HMI tags "IGG import"
   "RESET_STEP" : Bool = PLC RESET_STEP AT %M12.0, 1 s
   "Start Sequenc_DB_Post Purge Time Sec" : Int AT %DB1.DBW0
   "Tank Activated Port 10" : Int AT %DB1.DBW0
   "Tank Activated Port 2" : Int AT %DB1.DBW0
   "Tank Activated Port 3" : Int AT %DB1.DBW0
   "Tank Activated Port 4" : Int AT %DB1.DBW0
   "Tank Activated Port 5" : Int AT %DB1.DBW0
   "Tank Activated Port 6" : Int AT %DB1.DBW0
   "Tank Activated Port 7" : Int AT %DB1.DBW0
   "Tank Activated Port 8" : Int AT %DB1.DBW0
   "Tank Activated Port 9" : Int AT %DB1.DBW0
   "Tank Activated Star 10" : Int AT %DB1.DBW0
   "Tank Activated Star 2" : Int AT %DB1.DBW0
   "Tank Activated Star 3" : Int AT %DB1.DBW0
   "Tank Activated Star 4" : Int AT %DB1.DBW0
   "Tank Activated Star 5" : Int AT %DB1.DBW0
   "Tank Activated Star 6" : Int AT %DB1.DBW0
   "Tank Activated Star 7" : Int AT %DB1.DBW0
   "Tank Activated Star 8" : Int AT %DB1.DBW0
   "Tank Activated Star 9" : Int AT %DB1.DBW0
   "user_group" : Int AT %DB1.DBW0
   "2084_Setpoints_FIT417_HiHi" : Real = PLC "2084_Setpoints".FIT417_HiHi, 1 s
   "2086_Times_Tank Alarm Reset Time" : Time = PLC "2086_Times"."Tank Alarm Reset Time", 1 s
   "2084_Setpoints_FIT417_LoLo" : Real = PLC "2084_Setpoints".FIT417_LoLo, 1 s
   "2086_Times_Alarm Enable Delay" : Time = PLC "2086_Times"."Alarm Enable Delay", 1 s
   "2084_Setpoints_FIT417_Lo" : Real = PLC "2084_Setpoints".FIT417_Lo, 1 s
   "2084_Setpoints_FIT419_Lo" : Real = PLC "2084_Setpoints".FIT419_Lo, 1 s
   "2084_Setpoints_FIT417_Hi" : Real = PLC "2084_Setpoints".FIT417_Hi, 1 s
   "LT422 FPT  TANK LEVEL ALARM_LOW LEVEL VALUE (L)" : Real = PLC "LT422 FPT  TANK LEVEL ALARM"."LOW LEVEL VALUE (L)" AT %DB2226.DBD26, 1 s
   "2084_Setpoints_FIT419_LoLo" : Real = PLC "2084_Setpoints".FIT419_LoLo, 1 s
   "LT422 FPT  TANK LEVEL ALARM_ALARM L" : Bool = PLC "LT422 FPT  TANK LEVEL ALARM"."ALARM L" AT %DB2226.DBX48.2, 1 s
   "20_TANKS_IP_DATA_RIO_03_FIRST_TANK_O2_MONITOR" : Real = PLC "20_TANKS_IP_DATA".RIO_03.FIRST_TANK.O2_MONITOR, 1 s
   "20_TANKS_IP_DATA_RIO_07_FIRST_TANK_DECK_IG_PRESS" : Real = PLC "20_TANKS_IP_DATA".RIO_07.FIRST_TANK.DECK_IG_PRESS, 1 s
   "2062_Warning_Data_Alarm Tank FPT" : Bool = PLC "2062_Warning_Data"."Alarm Tank FPT" AT %DB2062.DBX22.1, 1 s
   "2084_Setpoints_LT421_Hi" : Real = PLC "2084_Setpoints".LT421_Hi, 1 s
   "2084_Setpoints_TX426 Port PH Lo" : Real = PLC "2084_Setpoints"."TX426 Port PH Lo", 1 s
   "2084_Setpoints_TX426 Port PH High" : Real = PLC "2084_Setpoints"."TX426 Port PH High", 1 s
   "2084_Setpoints_TX428 Port DO Lo" : Real = PLC "2084_Setpoints"."TX428 Port DO Lo", 1 s
   "2084_Setpoints_TX428 Port DO High" : Real = PLC "2084_Setpoints"."TX428 Port DO High", 1 s
   "2084_Setpoints_LT421_Lo" : Real = PLC "2084_Setpoints".LT421_Lo, 1 s
   "2084_Setpoints_FIT419_HiHi" : Real = PLC "2084_Setpoints".FIT419_HiHi, 1 s
   "2084_Setpoints_FIT419_Hi" : Real = PLC "2084_Setpoints".FIT419_Hi, 1 s
   "2084_Setpoints_TX425 Star PH Lo" : Real = PLC "2084_Setpoints"."TX425 Star PH Lo", 1 s
   "2084_Setpoints_TX425 Star PH High" : Real = PLC "2084_Setpoints"."TX425 Star PH High", 1 s
   "2084_Setpoints_TX427 Star DO Lo" : Real = PLC "2084_Setpoints"."TX427 Star DO Lo", 1 s
   "2084_Setpoints_TX427 Star DO High" : Real = PLC "2084_Setpoints"."TX427 Star DO High", 1 s
   "2084_Setpoints_Conf O2 Level Lo" : Real = PLC "2084_Setpoints"."Conf O2 Level Lo", 1 s
   "2084_Setpoints_Conf O2 Level Lo Lo" : Real = PLC "2084_Setpoints"."Conf O2 Level Lo Lo", 1 s
   "20_TANKS_IP_DATA_RIO_03_FIRST_TANK_DECK_IG_PRESS" : Real = PLC "20_TANKS_IP_DATA".RIO_03.FIRST_TANK.DECK_IG_PRESS, 1 s
   "20_TANKS_IP_DATA_RIO_01_THIRD_TANK_O2_MONITOR" : Real = PLC "20_TANKS_IP_DATA".RIO_01.THIRD_TANK.O2_MONITOR, 1 s
   "20_TANKS_IP_DATA_RIO_01_THIRD_TANK_DECK_IG_PRESS" : Real = PLC "20_TANKS_IP_DATA".RIO_01.THIRD_TANK.DECK_IG_PRESS, 1 s
   "20_TANKS_IP_DATA_RIO_01_FIRST_TANK_DECK_IG_PRESS" : Real = PLC "20_TANKS_IP_DATA".RIO_01.FIRST_TANK.DECK_IG_PRESS, 1 s
   "20_TANKS_IP_DATA_RIO_01_FIRST_TANK_O2_MONITOR" : Real = PLC "20_TANKS_IP_DATA".RIO_01.FIRST_TANK.O2_MONITOR, 1 s
   "20_TANKS_IP_DATA_RIO_04_FIRST_TANK_DECK_IG_PRESS" : Real = PLC "20_TANKS_IP_DATA".RIO_04.FIRST_TANK.DECK_IG_PRESS, 1 s
   "20_TANKS_IP_DATA_RIO_04_FIRST_TANK_O2_MONITOR" : Real = PLC "20_TANKS_IP_DATA".RIO_04.FIRST_TANK.O2_MONITOR, 1 s
   "20_TANKS_IP_DATA_RIO_04_SECOND_TANK_O2_MONITOR" : Real = PLC "20_TANKS_IP_DATA".RIO_04.SECOND_TANK.O2_MONITOR, 1 s
   "20_TANKS_IP_DATA_RIO_05_FIRST_TANK_DECK_IG_PRESS" : Real = PLC "20_TANKS_IP_DATA".RIO_05.FIRST_TANK.DECK_IG_PRESS, 1 s
   "20_TANKS_IP_DATA_RIO_05_FIRST_TANK_O2_MONITOR" : Real = PLC "20_TANKS_IP_DATA".RIO_05.FIRST_TANK.O2_MONITOR, 1 s
   "20_TANKS_IP_DATA_RIO_05_SECOND_TANK_O2_MONITOR" : Real = PLC "20_TANKS_IP_DATA".RIO_05.SECOND_TANK.O2_MONITOR, 1 s
   "20_TANKS_IP_DATA_RIO_06_FIRST_TANK_DECK_IG_PRESS" : Real = PLC "20_TANKS_IP_DATA".RIO_06.FIRST_TANK.DECK_IG_PRESS, 1 s
   "20_TANKS_IP_DATA_RIO_06_FIRST_TANK_O2_MONITOR" : Real = PLC "20_TANKS_IP_DATA".RIO_06.FIRST_TANK.O2_MONITOR, 1 s
   "20_TANKS_IP_DATA_RIO_07_FIRST_TANK_O2_MONITOR" : Real = PLC "20_TANKS_IP_DATA".RIO_07.FIRST_TANK.O2_MONITOR, 1 s
   "20_TANKS_IP_DATA_RIO_03_SECOND_TANK_O2_MONITOR" : Real = PLC "20_TANKS_IP_DATA".RIO_03.SECOND_TANK.O2_MONITOR, 1 s
   "2062_Warning_Data_Water Level Override FPT" : Bool = PLC "2062_Warning_Data"."Water Level Override FPT" AT %DB2062.DBX360.0, 1 s
   "Tank 3P Tank Vent Valve 2 Feedback - Closed" : Bool = PLC "Tank 3P Tank Vent Valve 2 Feedback - Closed" AT %I27.5, 1 s
   "2062_Warning_Data_Alarm Tank P1" : Bool = PLC "2062_Warning_Data"."Alarm Tank P1" AT %DB2062.DBX22.2, 1 s
   "Tank 2S Tank Vent Valve 2 Feedback - Opened" : Bool = PLC "Tank 2S Tank Vent Valve 2 Feedback - Opened" AT %I18.4, 1 s
   "Tank 2S Tank Vent Valve 1 Feedback - Closed" : Bool = PLC "Tank 2S Tank Vent Valve 1 Feedback - Closed" AT %I18.3, 1 s
   "Tank 2S Tank Vent Valve 1 Feedback - Opened" : Bool = PLC "Tank 2S Tank Vent Valve 1 Feedback - Opened" AT %I18.2, 1 s
   "Tank 2S GTT Isolation Valve Feedback - Closed" : Bool = PLC "Tank 2S GTT Isolation Valve Feedback - Closed" AT %I18.1, 1 s
   "Tank 2S GTT Isolation Valve Feedback - Opened" : Bool = PLC "Tank 2S GTT Isolation Valve Feedback - Opened" AT %I18.0, 1 s
   "RIO2_SPR_DI_15_7" : Bool = PLC RIO2_SPR_DI_15_7 AT %I15.7, 1 s
   "RIO2_SPR_DI_15_6" : Bool = PLC RIO2_SPR_DI_15_6 AT %I15.6, 1 s
   "Tank 2P Tank Vent Valve 2 Feedback - Closed" : Bool = PLC "20_TANKS_IP_DATA".RIO_05.FIRST_TANK.BWT_DO AT %I15.5, 1 s
   "Tank 2P Tank Vent Valve 2 Feedback - Opened" : Bool = PLC "Tank 2P Tank Vent Valve 2 Feedback - Opened" AT %I15.4, 1 s
   "Tank 2P Tank Vent Valve 1 Feedback - Closed" : Bool = PLC "Tank 2P Tank Vent Valve 1 Feedback - Closed" AT %I15.3, 1 s
   "Tank 2P Tank Vent Valve 1 Feedback - Opened" : Bool = PLC "Tank 2P Tank Vent Valve 1 Feedback - Opened" AT %I15.2, 1 s
   "Tank 2S Tank Vent Valve 2 Feedback - Closed" : Bool = PLC "Tank 2S Tank Vent Valve 2 Feedback - Closed" AT %I18.5, 1 s
   "Tank 2P GTT Isolation Valve Feedback - Closed" : Bool = PLC "Tank 2P GTT Isolation Valve Feedback - Closed" AT %I15.1, 1 s
   "RIO1_SPR_DI_9_7" : Bool = PLC RIO1_SPR_DI_9_7 AT %I9.7, 1 s
   "RIO1_SPR_DI_9_6" : Bool = PLC RIO1_SPR_DI_9_6 AT %I9.6, 1 s
   "RIO1_SPR_DI_9_5" : Bool = PLC RIO1_SPR_DI_9_5 AT %I9.5, 1 s
   "RIO1_SPR_DI_9_4" : Bool = PLC RIO1_SPR_DI_9_4 AT %I9.4, 1 s
   "Tank 1S BWT Level High High Switch" : Bool = PLC "Tank 1S BWT Level High High Switch" AT %I9.3, 1 s
   "Tank 1P BWT Level High High Switch" : Bool = PLC "Tank 1P BWT Level High High Switch" AT %I9.2, 1 s
   "RIO1 Tanks Pressure Switch Hi Hi" : Bool = PLC "RIO1 Tanks Pressure Switch Hi Hi" AT %I9.1, 1 s
   "FPT BWT Level High High Switch" : Bool = PLC "FPT BWT Level High High Switch" AT %I9.0, 1 s
   "RIO1_SPR_DI_6_7" : Bool = PLC RIO1_SPR_DI_6_7 AT %I6.7, 1 s
   "RIO1_SPR_DI_6_6" : Bool = PLC RIO1_SPR_DI_6_6 AT %I6.6, 1 s
   "Tank 1S Tank Vent Valve 2 Feedback - Closed" : Bool = PLC "Tank 1S Tank Vent Valve 2 Feedback - Closed" AT %I6.5, 1 s
   "Tank 2P GTT Isolation Valve Feedback - Opened" : Bool = PLC "Tank 2P GTT Isolation Valve Feedback - Opened" AT %I15.0, 1 s
   "RIO2_SPR_DI_18_6" : Bool = PLC RIO2_SPR_DI_18_6 AT %I18.6, 1 s
   "RIO2_SPR_DI_18_7" : Bool = PLC RIO2_SPR_DI_18_7 AT %I18.7, 1 s
   "Tank 2P BWT Level High High Switch" : Bool = PLC "Tank 2P BWT Level High High Switch" AT %I21.0, 1 s
   "RIO3 Tanks Pressure Switch Hi Hi" : Bool = PLC "RIO3 Tanks Pressure Switch Hi Hi" AT %I33.1, 1 s
   "Tank 3P BWT Level High High Switch" : Bool = PLC "Tank 3P BWT Level High High Switch" AT %I33.0, 1 s
   "RIO3_SPR_DI_30_7" : Bool = PLC RIO3_SPR_DI_30_7 AT %I30.7, 1 s
   "RIO3_SPR_DI_30_6" : Bool = PLC RIO3_SPR_DI_30_6 AT %I30.6, 1 s
   "Tank 3S Tank Vent Valve 2 Feedback - Closed" : Bool = PLC "Tank 3S Tank Vent Valve 2 Feedback - Closed" AT %I30.5, 1 s
   "Tank 3S Tank Vent Valve 2 Feedback - Opened" : Bool = PLC "Tank 3S Tank Vent Valve 2 Feedback - Opened" AT %I30.4, 1 s
   "Tank 3S Tank Vent Valve 1 Feedback - Closed" : Bool = PLC "Tank 3S Tank Vent Valve 1 Feedback - Closed" AT %I30.3, 1 s
   "Tank 3S Tank Vent Valve 1 Feedback - Opened" : Bool = PLC "Tank 3S Tank Vent Valve 1 Feedback - Opened" AT %I30.2, 1 s
   "Tank 3S GTT Isolation Valve Feedback - Closed" : Bool = PLC "Tank 3S GTT Isolation Valve Feedback - Closed" AT %I30.1, 1 s
   "Tank 3S GTT Isolation Valve Feedback - Opened" : Bool = PLC "Tank 3S GTT Isolation Valve Feedback - Opened" AT %I30.0, 1 s
   "RIO3_SPR_DI_27_7" : Bool = PLC RIO3_SPR_DI_27_7 AT %I27.7, 1 s
   "RIO3_SPR_DI_27_6" : Bool = PLC "63_Safety System Interlock_IDB"."Lockout Healthy" AT %I27.6, 1 s
   "504_Tank Grouping_DB2020_Diff Time Remain" : DInt = PLC "504_Tank Grouping_DB2020"."Diff Time Remain", 1 s
   "Tank 3P Tank Vent Valve 2 Feedback - Opened" : Bool = PLC "Tank 3P Tank Vent Valve 2 Feedback - Opened" AT %I27.4, 1 s
   "Tank 3P Tank Vent Valve 1 Feedback - Closed" : Bool = PLC "Tank 3P Tank Vent Valve 1 Feedback - Closed" AT %I27.3, 1 s
   "Tank 3P Tank Vent Valve 1 Feedback - Opened" : Bool = PLC "Tank 3P Tank Vent Valve 1 Feedback - Opened" AT %I27.2, 1 s
   "Tank 3P GTT Isolation Valve Feedback - Closed" : Bool = PLC "Tank 3P GTT Isolation Valve Feedback - Closed" AT %I27.1, 1 s
   "Tank 3P GTT Isolation Valve Feedback - Opened" : Bool = PLC "Tank 3P GTT Isolation Valve Feedback - Opened" AT %I27.0, 1 s
   "RIO2_SPR_DI_21_7" : Bool = PLC RIO2_SPR_DI_21_7 AT %I21.7, 1 s
   "RIO2_SPR_DI_21_6" : Bool = PLC RIO2_SPR_DI_21_6 AT %I21.6, 1 s
   "RIO2_SPR_DI_21_5" : Bool = PLC RIO2_SPR_DI_21_5 AT %I21.5, 1 s
   "RIO2_SPR_DI_21_4" : Bool = PLC RIO2_SPR_DI_21_4 AT %I21.4, 1 s
   "RIO2_SPR_DI_21_3" : Bool = PLC RIO2_SPR_DI_21_3 AT %I21.3, 1 s
   "Tank 2S BWT Level High High Switch" : Bool = PLC "Tank 2S BWT Level High High Switch" AT %I21.2, 1 s
   "RIO2 Tanks Pressure Switch Hi Hi" : Bool = PLC "RIO2 Tanks Pressure Switch Hi Hi" AT %I21.1, 1 s
   "Tank 1S Tank Vent Valve 2 Feedback - Opened" : Bool = PLC "Tank 1S Tank Vent Valve 2 Feedback - Opened" AT %I6.4, 1 s
   "Tank 1S Tank Vent Valve 1 Feedback - Closed" : Bool = PLC "Tank 1S Tank Vent Valve 1 Feedback - Closed" AT %I6.3, 1 s
   "Tank 1S Tank Vent Valve 1 Feedback - Opened" : Bool = PLC "Tank 1S Tank Vent Valve 1 Feedback - Opened" AT %I6.2, 1 s
   "Tank 1S GTT Isolation Valve Feedback - Closed" : Bool = PLC "Tank 1S GTT Isolation Valve Feedback - Closed" AT %I6.1, 1 s
   "2062_Warning_Data_Water Level Override 5P" : Bool = PLC "2062_Warning_Data"."Water Level Override 5P" AT %DB2062.DBX361.1, 1 s
   "2062_Warning_Data_Alarm Tank P5" : Bool = PLC "2062_Warning_Data"."Alarm Tank P5" AT %DB2062.DBX23.2, 1 s
   "LT422 5P  TANK LEVEL ALARM_ALARM L" : Bool = PLC "LT422 5P  TANK LEVEL ALARM"."ALARM L" AT %DB2235.DBX48.2, 1 s
   "2062_Warning_Data_Water Level Override 4S" : Bool = PLC "2062_Warning_Data"."Water Level Override 4S" AT %DB2062.DBX361.0, 1 s
   "2062_Warning_Data_Alarm Tank S4" : Bool = PLC "2062_Warning_Data"."Alarm Tank S4" AT %DB2062.DBX23.1, 1 s
   "LT421 4S  TANK LEVEL ALARM_ALARM L" : Bool = PLC "LT421 4S  TANK LEVEL ALARM"."ALARM L" AT %DB2234.DBX48.2, 1 s
   "2062_Warning_Data_Water Level Override 4P" : Bool = PLC "2062_Warning_Data"."Water Level Override 4P" AT %DB2062.DBX360.7, 1 s
   "2062_Warning_Data_Alarm Tank P4" : Bool = PLC "2062_Warning_Data"."Alarm Tank P4" AT %DB2062.DBX23.0, 1 s
   "LT422 4P  TANK LEVEL ALARM_ALARM L" : Bool = PLC "LT422 4P  TANK LEVEL ALARM"."ALARM L" AT %DB2233.DBX48.2, 1 s
   "2062_Warning_Data_Water Level Override 3S" : Bool = PLC "2062_Warning_Data"."Water Level Override 3S" AT %DB2062.DBX360.6, 1 s
   "2062_Warning_Data_Alarm Tank S3" : Bool = PLC "2062_Warning_Data"."Alarm Tank S3" AT %DB2062.DBX22.7, 1 s
   "LT421 3S  TANK LEVEL ALARM_ALARM L" : Bool = PLC "LT421 3S  TANK LEVEL ALARM"."ALARM L" AT %DB2232.DBX48.2, 1 s
   "2062_Warning_Data_Water Level Override 3P" : Bool = PLC "2062_Warning_Data"."Water Level Override 3P" AT %DB2062.DBX360.5, 1 s
   "2062_Warning_Data_Alarm Tank P3" : Bool = PLC "2062_Warning_Data"."Alarm Tank P3" AT %DB2062.DBX22.6, 1 s
   "LT422 3P  TANK LEVEL ALARM_ALARM L" : Bool = PLC "LT422 3P  TANK LEVEL ALARM"."ALARM L" AT %DB2231.DBX48.2, 1 s
   "2062_Warning_Data_Water Level Override 2S" : Bool = PLC "2062_Warning_Data"."Water Level Override 2S" AT %DB2062.DBX360.4, 1 s
   "2062_Warning_Data_Alarm Tank S2" : Bool = PLC "2062_Warning_Data"."Alarm Tank S2" AT %DB2062.DBX22.5, 1 s
   "LT421 2S  TANK LEVEL ALARM_ALARM L" : Bool = PLC "LT421 2S  TANK LEVEL ALARM"."ALARM L" AT %DB2230.DBX48.2, 1 s
   "2062_Warning_Data_Water Level Override 1S" : Bool = PLC "2062_Warning_Data"."Water Level Override 1S" AT %DB2062.DBX360.2, 1 s
   "2062_Warning_Data_Water Level Override 2P" : Bool = PLC "2062_Warning_Data"."Water Level Override 2P" AT %DB2062.DBX360.3, 1 s
   "2062_Warning_Data_Alarm Tank P2" : Bool = PLC "2062_Warning_Data"."Alarm Tank P2" AT %DB2062.DBX22.4, 1 s
   "FIT418_2P_ALM_ANALOG_DB_ALARM L" : Bool = PLC FIT418_2P_ALM_ANALOG_DB."ALARM L" AT %DB2064.DBX48.2, 1 s
   "2062_Warning_Data_Alarm Tank S1" : Bool = PLC "2062_Warning_Data"."Alarm Tank S1" AT %DB2062.DBX22.3, 1 s
   "LT421 1S  TANK LEVEL ALARM_ALARM L" : Bool = PLC "LT421 1S  TANK LEVEL ALARM"."ALARM L" AT %DB2228.DBX48.2, 1 s
   "2062_Warning_Data_Water Level Override 1P" : Bool = PLC "2062_Warning_Data"."Water Level Override 1P" AT %DB2062.DBX360.1, 1 s
   "LT421 5S  TANK LEVEL ALARM_ALARM L" : Bool = PLC "LT421 5S  TANK LEVEL ALARM"."ALARM L" AT %DB2236.DBX48.2, 1 s
   "LT422 1P  TANK LEVEL ALARM_ALARM L" : Bool = PLC "LT422 1P  TANK LEVEL ALARM"."ALARM L" AT %DB2227.DBX48.2, 1 s
   "2062_Warning_Data_Alarm Tank S5" : Bool = PLC "2062_Warning_Data"."Alarm Tank S5" AT %DB2062.DBX23.3, 1 s
   "LT422 6P  TANK LEVEL ALARM_ALARM L" : Bool = PLC "LT422 6P  TANK LEVEL ALARM"."ALARM L" AT %DB2237.DBX48.2, 1 s
   "Tank 1S GTT Isolation Valve Feedback - Opened" : Bool = PLC "Tank 1S GTT Isolation Valve Feedback - Opened" AT %I6.0, 1 s
   "RIO1_SPR_DI_3_7" : Bool = PLC RIO1_SPR_DI_3_7 AT %I3.7, 1 s
   "RIO1_SPR_DI_3_6" : Bool = PLC RIO1_SPR_DI_3_6 AT %I3.6, 1 s
   "Tank 1P Tank Vent Valve 2 Feedback - Closed" : Bool = PLC "Tank 1P Tank Vent Valve 2 Feedback - Closed" AT %I3.5, 1 s
   "Tank 1P Tank Vent Valve 2 Feedback - Opened" : Bool = PLC "Tank 1P Tank Vent Valve 2 Feedback - Opened" AT %I3.4, 1 s
   "Tank 1P Tank Vent Valve 1 Feedback - Closed" : Bool = PLC "Tank 1P Tank Vent Valve 1 Feedback - Closed" AT %I3.3, 1 s
   "Tank 1P Tank Vent Valve 1 Feedback - Opened" : Bool = PLC "Tank 1P Tank Vent Valve 1 Feedback - Opened" AT %I3.2, 1 s
   "Tank 1P GTT Isolation Valve Feedback - Closed" : Bool = PLC "Tank 1P GTT Isolation Valve Feedback - Closed" AT %I3.1, 1 s
   "Tank 1P GTT Isolation Valve Feedback - Opened" : Bool = PLC "Tank 1P GTT Isolation Valve Feedback - Opened" AT %I3.0, 1 s
   "RIO1_SPR_DI_0_7" : Bool = PLC RIO1_SPR_DI_0_7 AT %I0.7, 1 s
   "RIO1_SPR_DI_0_6" : Bool = PLC RIO1_SPR_DI_0_6 AT %I0.6, 1 s
   "FPT Tank Vent Valve 2 Feedback - Closed" : Bool = PLC "FPT Tank Vent Valve 2 Feedback - Closed" AT %I0.5, 1 s
   "FPT Tank Vent Valve 2 Feedback - Opened" : Bool = PLC "FPT Tank Vent Valve 2 Feedback - Opened" AT %I0.4, 1 s
   "FPT Tank Vent Valve 1 Feedback - Closed" : Bool = PLC "FPT Tank Vent Valve 1 Feedback - Closed" AT %I0.3, 1 s
   "FPT Tank Vent Valve 1 Feedback - Opened" : Bool = PLC "FPT Tank Vent Valve 1 Feedback - Opened" AT %I0.2, 1 s
   "FPT GTT Isolation Valve Feedback - Closed" : Bool = PLC "FPT GTT Isolation Valve Feedback - Closed" AT %I0.1, 1 s
   "FPT GTT Isolation Valve Feedback - Opened" : Bool = PLC "FPT GTT Isolation Valve Feedback - Opened" AT %I0.0, 1 s
   "2062_Warning_Data_Water Level Override APT" : Bool = PLC "2062_Warning_Data"."Water Level Override APT" AT %DB2062.DBX361.5, 1 s
   "2062_Warning_Data_Alarm Tank APT" : Bool = PLC "2062_Warning_Data"."Alarm Tank APT" AT %DB2062.DBX23.6, 1 s
   "LT422 APT  TANK LEVEL ALARM_ALARM L" : Bool = PLC "LT422 APT  TANK LEVEL ALARM"."ALARM L" AT %DB2239.DBX48.2, 1 s
   "2062_Warning_Data_Water Level Override 6S" : Bool = PLC "2062_Warning_Data"."Water Level Override 6S" AT %DB2062.DBX361.4, 1 s
   "2062_Warning_Data_Alarm Tank S6" : Bool = PLC "2062_Warning_Data"."Alarm Tank S6" AT %DB2062.DBX23.5, 1 s
   "LT421 6S  TANK LEVEL ALARM_ALARM L" : Bool = PLC "LT421 6S  TANK LEVEL ALARM"."ALARM L" AT %DB2238.DBX48.2, 1 s
   "2062_Warning_Data_Water Level Override 6P" : Bool = PLC "2062_Warning_Data"."Water Level Override 6P" AT %DB2062.DBX361.3, 1 s
   "2062_Warning_Data_Alarm Tank P6" : Bool = PLC "2062_Warning_Data"."Alarm Tank P6" AT %DB2062.DBX23.4, 1 s
   "2062_Warning_Data_Water Level Override 5S" : Bool = PLC "2062_Warning_Data"."Water Level Override 5S" AT %DB2062.DBX361.2, 1 s
   "504_Tank Grouping_DB2020_SetGroupSR" : Bool = PLC "504_Tank Grouping_DB2020".SetGroupSR, 1 s
   "20_TANKS_IP_DATA_RIO_06_SECOND_TANK_MBG_FLOW" : Real = PLC "20_TANKS_IP_DATA".RIO_06.SECOND_TANK.MBG_FLOW, 1 s
   "504_Tank Grouping_DB2020_Time Left Tank_Time Left Tank 14" : Real = PLC "504_Tank Grouping_DB2020"."Time Left Tank"."Time Left Tank 14", 1 s
   "20_TANKS_IP_DATA_RIO_01_THIRD_TANK_GTT_ISOL_VALVE_OPEN" : Bool = PLC "20_TANKS_IP_DATA".RIO_01.THIRD_TANK.GTT_ISOL_VALVE_OPEN, 1 s
   "20_TANKS_IP_DATA_RIO_01_THIRD_TANK_MBG_FLOW" : Real = PLC "20_TANKS_IP_DATA".RIO_01.THIRD_TANK.MBG_FLOW, 1 s
   "20_TANKS_IP_DATA_RIO_01_THIRD_TANK_USD_FLOW" : Real = PLC "20_TANKS_IP_DATA".RIO_01.THIRD_TANK.USD_FLOW, 1 s
   "504_Tank Grouping_DB2020_RUN TANK 3" : Bool = PLC "504_Tank Grouping_DB2020"."RUN TANK 3", 1 s
   "20_TANKS_IP_DATA_RIO_01_THIRD_TANK_BWT_LEVEL_HIHI" : Bool = PLC "20_TANKS_IP_DATA".RIO_01.THIRD_TANK.BWT_LEVEL_HIHI, 1 s
   "20_TANKS_IP_DATA_RIO_01_FIRST_TANK_GTT_ISOL_VALVE_CLSD" : Bool = PLC "20_TANKS_IP_DATA".RIO_01.FIRST_TANK.GTT_ISOL_VALVE_CLSD, 1 s
   "20_TANKS_IP_DATA_RIO_01_SECOND_TANK_GTT_ISOL_VALVE_CLSD" : Bool = PLC "20_TANKS_IP_DATA".RIO_01.SECOND_TANK.GTT_ISOL_VALVE_CLSD, 1 s
   "20_TANKS_IP_DATA_RIO_01_SECOND_TANK_GTT_ISOL_VALVE_OPEN" : Bool = PLC "20_TANKS_IP_DATA".RIO_01.SECOND_TANK.GTT_ISOL_VALVE_OPEN, 1 s
   "20_TANKS_IP_DATA_RIO_01_SECOND_TANK_MBG_FLOW" : Real = PLC "20_TANKS_IP_DATA".RIO_01.SECOND_TANK.MBG_FLOW, 1 s
   "20_TANKS_IP_DATA_RIO_01_SECOND_TANK_USD_FLOW" : Real = PLC "20_TANKS_IP_DATA".RIO_01.SECOND_TANK.USD_FLOW, 1 s
   "20_TANKS_IP_DATA_RIO_01_SECOND_TANK_BWT_LEVEL_HIHI" : Bool = PLC "20_TANKS_IP_DATA".RIO_01.SECOND_TANK.BWT_LEVEL_HIHI, 1 s
   "504_Tank Grouping_DB2020_RUN TANK 2" : Bool = PLC "504_Tank Grouping_DB2020"."RUN TANK 2", 1 s
   "504_Tank Grouping_DB2020_RUN TANK 1" : Bool = PLC "504_Tank Grouping_DB2020"."RUN TANK 1", 1 s
   "20_TANKS_IP_DATA_RIO_01_FIRST_TANK_GTT_ISOL_VALVE_OPEN" : Bool = PLC "20_TANKS_IP_DATA".RIO_01.FIRST_TANK.GTT_ISOL_VALVE_OPEN, 1 s
   "20_TANKS_IP_DATA_RIO_01_FIRST_TANK_USD_FLOW" : Real = PLC "20_TANKS_IP_DATA".RIO_01.FIRST_TANK.USD_FLOW, 1 s
   "20_TANKS_IP_DATA_RIO_01_FIRST_TANK_MBG_FLOW" : Real = PLC "20_TANKS_IP_DATA".RIO_01.FIRST_TANK.MBG_FLOW, 1 s
   "20_TANKS_IP_DATA_RIO_01_FIRST_TANK_BWT_LEVEL_HIHI" : Bool = PLC "20_TANKS_IP_DATA".RIO_01.FIRST_TANK.BWT_LEVEL_HIHI, 1 s
   "HMI Indication Logic_DB_Sequence Finished" : Bool = PLC "HMI Indication Logic_DB"."Sequence Finished", 1 s
   "51_SLAVE_STATUS_RUNNING" : Bool = PLC "51_SLAVE_STATUS".RUNNING AT %DB51.DBX4.2, 1 s
   "HMI Indication Logic_DB_Tank Selected" : Bool = PLC "HMI Indication Logic_DB"."Tank Selected", 1 s
   "HMI Indication Logic_DB_FA Mode Selected" : Bool = PLC "HMI Indication Logic_DB"."FA Mode Selected", 1 s
   "80_From_HMI_TIMER RST Supres" : Bool = PLC "80_From_HMI"."TIMER RST Supres", 1 s
   "504_Tank Grouping_DB2020_GROUP ACTIVE INT 7" : Bool = PLC "504_Tank Grouping_DB2020"."GROUP ACTIVE INT 7", 1 s
   "504_Tank Grouping_DB2020_GROUP ACTIVE INT 6" : Bool = PLC "504_Tank Grouping_DB2020"."GROUP ACTIVE INT 6", 1 s
   "504_Tank Grouping_DB2020_GROUP ACTIVE INT 5" : Bool = PLC "504_Tank Grouping_DB2020"."GROUP ACTIVE INT 5", 1 s
   "20_TANKS_IP_DATA_RIO_01_THIRD_TANK_GTT_ISOL_VALVE_CLSD" : Bool = PLC "20_TANKS_IP_DATA".RIO_01.THIRD_TANK.GTT_ISOL_VALVE_CLSD, 1 s
   "504_Tank Grouping_DB2020_GROUP ACTIVE INT 4" : Bool = PLC "504_Tank Grouping_DB2020"."GROUP ACTIVE INT 4", 1 s
   "504_Tank Grouping_DB2020_RUN TANK 4" : Bool = PLC "504_Tank Grouping_DB2020"."RUN TANK 4", 1 s
   "20_TANKS_IP_DATA_RIO_03_FIRST_TANK_MBG_FLOW" : Real = PLC "20_TANKS_IP_DATA".RIO_03.FIRST_TANK.MBG_FLOW, 1 s
   "20_TANKS_IP_DATA_RIO_05_FIRST_TANK_GTT_ISOL_VALVE_CLSD" : Bool = PLC "20_TANKS_IP_DATA".RIO_05.FIRST_TANK.GTT_ISOL_VALVE_CLSD, 1 s
   "20_TANKS_IP_DATA_RIO_05_FIRST_TANK_GTT_ISOL_VALVE_OPEN" : Bool = PLC "20_TANKS_IP_DATA".RIO_05.FIRST_TANK.GTT_ISOL_VALVE_OPEN, 1 s
   "20_TANKS_IP_DATA_RIO_05_FIRST_TANK_USD_FLOW" : Real = PLC "20_TANKS_IP_DATA".RIO_05.FIRST_TANK.USD_FLOW, 1 s
   "20_TANKS_IP_DATA_RIO_05_FIRST_TANK_MBG_FLOW" : Real = PLC "20_TANKS_IP_DATA".RIO_05.FIRST_TANK.MBG_FLOW, 1 s
   "20_TANKS_IP_DATA_RIO_05_FIRST_TANK_BWT_LEVEL_HIHI" : Bool = PLC "20_TANKS_IP_DATA".RIO_05.FIRST_TANK.BWT_LEVEL_HIHI, 1 s
   "20_TANKS_IP_DATA_RIO_04_SECOND_TANK_GTT_ISOL_VALVE_CLSD" : Bool = PLC "20_TANKS_IP_DATA".RIO_04.SECOND_TANK.GTT_ISOL_VALVE_CLSD, 1 s
   "20_TANKS_IP_DATA_RIO_04_SECOND_TANK_GTT_ISOL_VALVE_OPEN" : Bool = PLC "20_TANKS_IP_DATA".RIO_04.SECOND_TANK.GTT_ISOL_VALVE_OPEN, 1 s
   "20_TANKS_IP_DATA_RIO_04_SECOND_TANK_MBG_FLOW" : Real = PLC "20_TANKS_IP_DATA".RIO_04.SECOND_TANK.MBG_FLOW, 1 s
   "20_TANKS_IP_DATA_RIO_04_SECOND_TANK_USD_FLOW" : Real = PLC "20_TANKS_IP_DATA".RIO_04.SECOND_TANK.USD_FLOW, 1 s
   "20_TANKS_IP_DATA_RIO_04_SECOND_TANK_BWT_LEVEL_HIHI" : Bool = PLC "20_TANKS_IP_DATA".RIO_04.SECOND_TANK.BWT_LEVEL_HIHI, 1 s
   "20_TANKS_IP_DATA_RIO_04_FIRST_TANK_GTT_ISOL_VALVE_CLSD" : Bool = PLC "20_TANKS_IP_DATA".RIO_04.FIRST_TANK.GTT_ISOL_VALVE_CLSD, 1 s
   "20_TANKS_IP_DATA_RIO_04_FIRST_TANK_GTT_ISOL_VALVE_OPEN" : Bool = PLC "20_TANKS_IP_DATA".RIO_04.FIRST_TANK.GTT_ISOL_VALVE_OPEN, 1 s
   "20_TANKS_IP_DATA_RIO_04_FIRST_TANK_MBG_FLOW" : Real = PLC "20_TANKS_IP_DATA".RIO_04.FIRST_TANK.MBG_FLOW, 1 s
   "20_TANKS_IP_DATA_RIO_04_FIRST_TANK_USD_FLOW" : Real = PLC "20_TANKS_IP_DATA".RIO_04.FIRST_TANK.USD_FLOW, 1 s
   "20_TANKS_IP_DATA_RIO_04_FIRST_TANK_BWT_LEVEL_HIHI" : Bool = PLC "20_TANKS_IP_DATA".RIO_04.FIRST_TANK.BWT_LEVEL_HIHI, 1 s
   "20_TANKS_IP_DATA_RIO_03_SECOND_TANK_GTT_ISOL_VALVE_CLSD" : Bool = PLC "20_TANKS_IP_DATA".RIO_03.SECOND_TANK.GTT_ISOL_VALVE_CLSD, 1 s
   "20_TANKS_IP_DATA_RIO_03_SECOND_TANK_GTT_ISOL_VALVE_OPEN" : Bool = PLC "20_TANKS_IP_DATA".RIO_03.SECOND_TANK.GTT_ISOL_VALVE_OPEN, 1 s
   "20_TANKS_IP_DATA_RIO_03_SECOND_TANK_MBG_FLOW" : Real = PLC "20_TANKS_IP_DATA".RIO_03.SECOND_TANK.MBG_FLOW, 1 s
   "20_TANKS_IP_DATA_RIO_03_SECOND_TANK_USD_FLOW" : Real = PLC "20_TANKS_IP_DATA".RIO_03.SECOND_TANK.USD_FLOW, 1 s
   "504_Tank Grouping_DB2020_RUN TANK 7" : Bool = PLC "504_Tank Grouping_DB2020"."RUN TANK 7", 1 s
   "20_TANKS_IP_DATA_RIO_03_SECOND_TANK_BWT_LEVEL_HIHI" : Bool = PLC "20_TANKS_IP_DATA".RIO_03.SECOND_TANK.BWT_LEVEL_HIHI, 1 s
   "20_TANKS_IP_DATA_RIO_03_FIRST_TANK_GTT_ISOL_VALVE_CLSD" : Bool = PLC "20_TANKS_IP_DATA".RIO_03.FIRST_TANK.GTT_ISOL_VALVE_CLSD, 1 s
   "20_TANKS_IP_DATA_RIO_03_FIRST_TANK_GTT_ISOL_VALVE_OPEN" : Bool = PLC "20_TANKS_IP_DATA".RIO_03.FIRST_TANK.GTT_ISOL_VALVE_OPEN, 1 s
   "20_TANKS_IP_DATA_RIO_03_FIRST_TANK_BWT_LEVEL_HIHI" : Bool = PLC "20_TANKS_IP_DATA".RIO_03.FIRST_TANK.BWT_LEVEL_HIHI, 1 s
   "20_TANKS_IP_DATA_RIO_03_FIRST_TANK_USD_FLOW" : Real = PLC "20_TANKS_IP_DATA".RIO_03.FIRST_TANK.USD_FLOW, 1 s
   "504_Tank Grouping_DB2020_RUN TANK 5" : Bool = PLC "504_Tank Grouping_DB2020"."RUN TANK 5", 1 s
   "504_Tank Grouping_DB2020_GROUP ACTIVE INT 3" : Bool = PLC "504_Tank Grouping_DB2020"."GROUP ACTIVE INT 3", 1 s
   "504_Tank Grouping_DB2020_GROUP ACTIVE INT 2" : Bool = PLC "504_Tank Grouping_DB2020"."GROUP ACTIVE INT 2", 1 s
   "504_Tank Grouping_DB2020_GROUP ACTIVE INT 1" : Bool = PLC "504_Tank Grouping_DB2020"."GROUP ACTIVE INT 1", 1 s
   "PGC_COMMISSION_MODE_DB_Drive Popup" : Bool = PLC PGC_COMMISSION_MODE_DB."Drive Popup", 500 ms
      on ChangeValue: "PGCCommissioning"()
   "PGC_COMMISSION_MODE_DB_Active" : Bool = PLC PGC_COMMISSION_MODE_DB.Active, 1 s
   "PGC_COMMISSION_MODE_DB_Button Control" : Int = PLC PGC_COMMISSION_MODE_DB."Button Control", 1 s
   "PGC_COMMISSION_MODE_DB_Setpoint" : Real = PLC PGC_COMMISSION_MODE_DB.Setpoint, 1 s
   "2102_TIME_CALCS_DB_Time_To_Treatment" : Int = PLC "2102_TIME_CALCS_DB".Time_To_Treatment, 1 s
   "2102_TIME_CALCS_DB_Voyage_TIME_remaining_h" : Int = PLC "2102_TIME_CALCS_DB".Voyage_TIME_remaining_h, 1 s
   "2102_TIME_CALCS_DB_Voyage_TIME_remaining_m" : Int = PLC "2102_TIME_CALCS_DB".Voyage_TIME_remaining_m, 1 s
   "2086_Times_PS436 Alarm Delay" : Time = PLC "2086_Times"."PS436 Alarm Delay", 1 s
   "2086_Times_LS425 Star Alarm Delay" : Time = PLC "2086_Times"."LS425 Star Alarm Delay", 1 s
   "2086_Times_LS425 Port Alarm Delay" : Time = PLC "2086_Times"."LS425 Port Alarm Delay", 1 s
   "2086_Times_PIT424 Alarm Delay" : Time = PLC "2086_Times"."PIT424 Alarm Delay", 1 s
   "2086_Times_PT415 Alarm Delay" : Time = PLC "2086_Times"."PT415 Alarm Delay", 1 s
   "2086_Times_FIT419STAR Alarm Delay" : Time = PLC "2086_Times"."FIT419STAR Alarm Delay", 1 s
   "2086_Times_FIT417STAR Alarm Delay" : Time = PLC "2086_Times"."FIT417STAR Alarm Delay", 1 s
   "2086_Times_FIT420PORT Alarm Delay" : Time = PLC "2086_Times"."FIT420PORT Alarm Delay", 1 s
   "2086_Times_FIT418PORT Alarm Delay" : Time = PLC "2086_Times"."FIT418PORT Alarm Delay", 1 s
   "2086_Times_TT426_STAR_Alarm Delay" : Time = PLC "2086_Times"."TT426_STAR_Alarm Delay", 1 s
   "2086_Times_TT426_PORT_Alarm Delay" : Time = PLC "2086_Times"."TT426_PORT_Alarm Delay", 1 s
   "84_Setpoints_LIT304_Refill_Target_Low" : Real = PLC "84_Setpoints".LIT304_Refill_Target_Low, 1 s
   "84_Setpoints_LIT304_InitialFill_Target_Low" : Real = PLC "84_Setpoints".LIT304_InitialFill_Target_Low, 1 s
   "2102_TIME_CALCS_DB_PRE-DWEL MINS REMNG" : Int = PLC "2102_TIME_CALCS_DB"."PRE-DWEL MINS REMNG", 1 s
   "21_FLOW_PRESSURE_SETPOINT_FIT_419_PRESSURE_SETPOINT" : Real = PLC "21_FLOW_PRESSURE_SETPOINT".FIT_419_PRESSURE_SETPOINT, 1 s
   "21_FLOW_PRESSURE_SETPOINT_FIT_420_PRESSURE_SETPOINT" : Real = PLC "21_FLOW_PRESSURE_SETPOINT".FIT_420_PRESSURE_SETPOINT, 1 s
   "2102_TIME_CALCS_DB_Voyage_TIME_hours" : Int = PLC "2102_TIME_CALCS_DB".Voyage_TIME_hours, 1 s
   "2115_VOYAGE_TIME_DAYS_VOYAGE_DAYS" : Real = PLC "80_From_HMI".MAN_DQ_1_3, 1 s
   "504_Tank Grouping_DB2020_GROUP SET" : Int = PLC "504_Tank Grouping_DB2020"."GROUP SET", 1 s
   "504_Tank Grouping_DB2020_GROUP ACTIV 7" : Bool = PLC "504_Tank Grouping_DB2020"."GROUP ACTIV 7", 1 s
   "504_Tank Grouping_DB2020_GROUP ACTIV 6" : Bool = PLC "504_Tank Grouping_DB2020"."GROUP ACTIV 6", 1 s
   "504_Tank Grouping_DB2020_GROUP ACTIV 5" : Bool = PLC "504_Tank Grouping_DB2020"."GROUP ACTIV 5", 1 s
   "504_Tank Grouping_DB2020_GROUP ACTIV 4" : Bool = PLC "504_Tank Grouping_DB2020"."GROUP ACTIV 4", 1 s
   "504_Tank Grouping_DB2020_GROUP ACTIV 3" : Bool = PLC "504_Tank Grouping_DB2020"."GROUP ACTIV 3", 1 s
   "504_Tank Grouping_DB2020_GROUP ACTIV 2" : Bool = PLC "504_Tank Grouping_DB2020"."GROUP ACTIV 2", 1 s
   "504_Tank Grouping_DB2020_GROUP ACTIV 1" : Bool = PLC "504_Tank Grouping_DB2020"."GROUP ACTIV 1", 1 s
   "504_Tank Grouping_DB2020_GROUP of TANK 14" : Int = PLC "504_Tank Grouping_DB2020"."GROUP of TANK 14", 1 s
   "504_Tank Grouping_DB2020_GROUP of TANK 13" : Int = PLC "504_Tank Grouping_DB2020"."GROUP of TANK 13", 1 s
   "504_Tank Grouping_DB2020_GROUP of TANK 12" : Int = PLC "504_Tank Grouping_DB2020"."GROUP of TANK 12", 1 s
   "504_Tank Grouping_DB2020_GROUP of TANK 11" : Int = PLC "504_Tank Grouping_DB2020"."GROUP of TANK 11", 1 s
   "20_TANKS_IP_DATA_RIO_05_SECOND_TANK_BWT_LEVEL_HIHI" : Bool = PLC "20_TANKS_IP_DATA".RIO_05.SECOND_TANK.BWT_LEVEL_HIHI, 1 s
   "504_Tank Grouping_DB2020_GROUP of TANK 10" : Int = PLC "504_Tank Grouping_DB2020"."GROUP of TANK 10", 1 s
   "504_Tank Grouping_DB2020_GROUP of TANK 8" : Int = PLC "504_Tank Grouping_DB2020"."GROUP of TANK 8", 1 s
   "504_Tank Grouping_DB2020_GROUP of TANK 7" : Int = PLC "504_Tank Grouping_DB2020"."GROUP of TANK 7", 1 s
   "504_Tank Grouping_DB2020_GROUP of TANK 6" : Int = PLC "504_Tank Grouping_DB2020"."GROUP of TANK 6", 1 s
   "504_Tank Grouping_DB2020_GROUP of TANK 5" : Int = PLC "504_Tank Grouping_DB2020"."GROUP of TANK 5", 1 s
   "504_Tank Grouping_DB2020_GROUP of TANK 4" : Int = PLC "504_Tank Grouping_DB2020"."GROUP of TANK 4", 1 s
   "504_Tank Grouping_DB2020_GROUP of TANK 3" : Int = PLC "504_Tank Grouping_DB2020"."GROUP of TANK 3", 1 s
   "504_Tank Grouping_DB2020_GROUP of TANK 2" : Int = PLC "504_Tank Grouping_DB2020"."GROUP of TANK 2", 1 s
   "504_Tank Grouping_DB2020_GROUP of TANK 1" : Int = PLC "504_Tank Grouping_DB2020"."GROUP of TANK 1", 1 s
   "504_Tank Grouping_DB2020_SetGroup" : Bool = PLC "504_Tank Grouping_DB2020".SetGroup, 1 s
   "2102_TIME_CALCS_DB_PHASE_DIFFERECE_MNS_REMNG_De-Ox" : Int = PLC "2102_TIME_CALCS_DB".PHASE_DIFFERECE_MNS_REMNG_De-Ox, 1 s
   "88_treatment_POP_UP_CNFRM" : Bool = PLC "88_treatment".POP_UP_CNFRM AT %DB1.DBX0.0, 1 s
   "88_treatment_POP_UP" : Bool = PLC "88_treatment".POP_UP AT %DB1.DBX0.0, 1 s
      on ChangeValue: "TreatmentdDailyChecks"()
   "504_Tank Grouping_DB2020_GROUP of TANK 9" : Int = PLC "504_Tank Grouping_DB2020"."GROUP of TANK 9", 1 s
   "504_Tank Grouping_DB2020_Time Left Tank_Time Left Tank 1" : Real = PLC "504_Tank Grouping_DB2020"."Time Left Tank"."Time Left Tank 1", 1 s
   "20_TANKS_IP_DATA_RIO_05_SECOND_TANK_USD_FLOW" : Real = PLC "20_TANKS_IP_DATA".RIO_05.SECOND_TANK.USD_FLOW, 1 s
   "20_TANKS_IP_DATA_RIO_05_SECOND_TANK_GTT_ISOL_VALVE_OPEN" : Bool = PLC "20_TANKS_IP_DATA".RIO_05.SECOND_TANK.GTT_ISOL_VALVE_OPEN, 1 s
   "20_TANKS_IP_DATA_RIO_06_FIRST_TANK_BWT_DO" : Real = PLC "2102_TIME_CALCS_DB".RE_OX_SP_MINS_RMNG, 1 s
   "20_TANKS_IP_DATA_RIO_06_FIRST_TANK_BWT_PH" : Real = PLC "20_TANKS_IP_DATA".RIO_06.FIRST_TANK.BWT_PH, 1 s
   "20_TANKS_IP_DATA_RIO_06_FIRST_TANK_BWT_LEVEL" : Real = PLC "20_TANKS_IP_DATA".RIO_06.FIRST_TANK.BWT_LEVEL, 1 s
   "20_TANKS_IP_DATA_RIO_06_FIRST_TANK_TANKS_PRESS" : Real = PLC "20_TANKS_IP_DATA".RIO_06.FIRST_TANK.TANKS_PRESS, 1 s
   "20_TANKS_IP_DATA_RIO_05_SECOND_TANK_BWT_TEMP" : Real = PLC "20_TANKS_IP_DATA".RIO_05.SECOND_TANK.BWT_TEMP, 1 s
   "20_TANKS_IP_DATA_RIO_05_SECOND_TANK_BWT_DO" : Real = PLC "20_TANKS_IP_DATA".RIO_05.SECOND_TANK.BWT_DO, 1 s
   "20_TANKS_IP_DATA_RIO_05_SECOND_TANK_BWT_PH" : Real = PLC "20_TANKS_IP_DATA".RIO_05.SECOND_TANK.BWT_PH, 1 s
   "20_TANKS_IP_DATA_RIO_05_SECOND_TANK_BWT_LEVEL" : Real = PLC "20_TANKS_IP_DATA".RIO_05.SECOND_TANK.BWT_LEVEL, 1 s
   "20_TANKS_IP_DATA_RIO_05_SECOND_TANK_TANKS_PRESS" : Real = PLC "20_TANKS_IP_DATA".RIO_05.SECOND_TANK.TANKS_PRESS, 1 s
   "504_Tank Grouping_DB2020_Tank10 Min Time_ET" : Time = PLC "504_Tank Grouping_DB2020"."Tank10 Min Time".ET, 1 s
   "20_TANKS_IP_DATA_RIO_05_FIRST_TANK_BWT_TEMP" : Real = PLC "20_TANKS_IP_DATA".RIO_05.FIRST_TANK.BWT_TEMP, 1 s
   "20_TANKS_IP_DATA_RIO_05_FIRST_TANK_BWT_DO" : Real = PLC "20_TANKS_IP_DATA".RIO_05.FIRST_TANK.BWT_DO, 1 s
   "20_TANKS_IP_DATA_RIO_05_FIRST_TANK_BWT_PH" : Real = PLC "20_TANKS_IP_DATA".RIO_05.FIRST_TANK.BWT_PH, 1 s
   "20_TANKS_IP_DATA_RIO_05_FIRST_TANK_BWT_LEVEL" : Real = PLC "20_TANKS_IP_DATA".RIO_05.FIRST_TANK.BWT_LEVEL, 1 s
   "20_TANKS_IP_DATA_RIO_05_FIRST_TANK_TANKS_PRESS" : Real = PLC "20_TANKS_IP_DATA".RIO_05.FIRST_TANK.TANKS_PRESS, 1 s
   "504_Tank Grouping_DB2020_Tank9 Min Time_ET" : Time = PLC "504_Tank Grouping_DB2020"."Tank9 Min Time".ET, 1 s
   "20_TANKS_IP_DATA_RIO_04_SECOND_TANK_BWT_TEMP" : Real = PLC "20_TANKS_IP_DATA".RIO_04.SECOND_TANK.BWT_TEMP, 1 s
   "20_TANKS_IP_DATA_RIO_04_SECOND_TANK_BWT_DO" : Real = PLC "20_TANKS_IP_DATA".RIO_04.SECOND_TANK.BWT_DO, 1 s
   "20_TANKS_IP_DATA_RIO_04_SECOND_TANK_BWT_PH" : Real = PLC "20_TANKS_IP_DATA".RIO_04.SECOND_TANK.BWT_PH, 1 s
   "20_TANKS_IP_DATA_RIO_04_SECOND_TANK_BWT_LEVEL" : Real = PLC "20_TANKS_IP_DATA".RIO_04.SECOND_TANK.BWT_LEVEL, 1 s
   "20_TANKS_IP_DATA_RIO_04_SECOND_TANK_TANKS_PRESS" : Real = PLC "20_TANKS_IP_DATA".RIO_04.SECOND_TANK.TANKS_PRESS, 1 s
   "504_Tank Grouping_DB2020_Tank8 Min Time_ET" : Time = PLC "504_Tank Grouping_DB2020"."Tank8 Min Time".ET, 1 s